screen "BWT Digital Inputs" 1280x800, template "Template"
   on GenerateScreen: "TitleUpdater"()
   TextField "Text field_37" at 16,52 size 263x26; Text 'BWT Control PLC (Rack 3)'
   TextField "Text field_38" at 16,122 size 55x22; Text 'I0.0'
   TextField "Text field_39" at 16,158 size 55x22; Text 'I0.1'
   TextField "Text field_40" at 16,194 size 55x22; Text 'I0.2'
   TextField "Text field_41" at 16,230 size 55x22; Text 'I0.3'
   TextField "Text field_42" at 16,265 size 55x22; Text 'I0.4'
   TextField "Text field_43" at 16,301 size 55x22; Text 'I0.5'
   TextField "Text field_44" at 16,337 size 55x22; Text 'I0.6'
   TextField "Text field_45" at 16,373 size 55x22; Text 'I0.7'
   Circle "Circle_33" at 76,122 size 20x20
      Appearance <- "10 DI_DATA_PS101"
   Circle "Circle_34" at 76,158 size 20x20
      Appearance <- "10 DI_DATA_E131_SHTDN"
   Circle "Circle_35" at 76,194 size 20x20
      Appearance <- "10 DI_DATA_R2_SPR_DI_0_2"
   Circle "Circle_36" at 76,230 size 20x20
      Appearance <- "10 DI_DATA_R2_SPR_DI_0_3"
   Circle "Circle_37" at 76,265 size 20x20
      Appearance <- "10 DI_DATA_X001_PWR_OK"
   Circle "Circle_38" at 76,301 size 20x20
      Appearance <- "10 DI_DATA_FD001_PWR_OK"
   Circle "Circle_39" at 76,337 size 20x20
      Appearance <- "10 DI_DATA_FD001_OK"
   Circle "Circle_40" at 76,373 size 20x20
      Appearance <- "103_Main_Burner_DB_DN_OK(1)"
   TextField "Text field_46" at 33,90 size 49x26; Text 'I0'
   TextField "Text field_47" at 16,441 size 55x22; Text 'I1.0'
   TextField "Text field_48" at 16,477 size 55x22; Text 'I1.1'
   TextField "Text field_49" at 16,513 size 55x22; Text 'I1.2'
   TextField "Text field_50" at 16,549 size 55x22; Text 'I1.3'
   TextField "Text field_51" at 16,584 size 55x22; Text 'I1.4'
   TextField "Text field_52" at 16,620 size 55x22; Text 'I1.5'
   TextField "Text field_53" at 16,656 size 55x22; Text 'I1.6'
   TextField "Text field_54" at 16,692 size 55x22; Text 'I1.7'
   Circle "Circle_41" at 76,441 size 20x20
      Appearance <- "10 DI_DATA_FS123"
   Circle "Circle_42" at 76,477 size 20x20
      Appearance <- "10 DI_DATA_FS115(1)"
   Circle "Circle_43" at 76,513 size 20x20
      Appearance <- "10 DI_DATA_FS320"
   Circle "Circle_44" at 76,549 size 20x20
      Appearance <- "10 DI_DATA_FS317"
   Circle "Circle_45" at 76,584 size 20x20
      Appearance <- "10 DI_DATA_P301_TRIPPED(1)"
   Circle "Circle_46" at 76,620 size 20x20
      Appearance <- "10 DI_DATA_P301_ENBLD"
   Circle "Circle_47" at 76,656 size 20x20
      Appearance <- "10 DI_DATA_R2_SPR_DI_1_6"
   Circle "Circle_48" at 76,692 size 20x20
      Appearance <- "10 DI_DATA_ESD_OK"
   TextField "Text field_55" at 33,409 size 49x26; Text 'I1'
   TextField "Text field_56" at 307,122 size 55x22; Text 'I2.0'
   TextField "Text field_57" at 307,158 size 55x22; Text 'I2.1'
   TextField "Text field_58" at 307,194 size 55x22; Text 'I2.2'
   TextField "Text field_59" at 307,230 size 55x22; Text 'I2.3'
   TextField "Text field_60" at 307,265 size 55x22; Text 'I2.4'
   TextField "Text field_61" at 307,301 size 55x22; Text 'I2.5'
   TextField "Text field_62" at 307,337 size 55x22; Text 'I2.6'
   TextField "Text field_63" at 307,373 size 55x22; Text 'I2.7'
   Circle "Circle_49" at 367,122 size 20x20
      Appearance <- "10 DI_DATA_E600_NOK"
   Circle "Circle_50" at 367,158 size 20x20
      Appearance <- "10 DI_DATA_E600_HIHI"
   Circle "Circle_51" at 367,194 size 20x20
      Appearance <- "10 DI_DATA_E600_LOLO"
   Circle "Circle_52" at 367,230 size 20x20
      Appearance <- "10 DI_DATA_E600_PWR_OK"
   Circle "Circle_53" at 367,265 size 20x20
      Appearance <- "10 DI_DATA_E700_PWR_OK"
   Circle "Circle_54" at 367,301 size 20x20
      Appearance <- "10 DI_DATA_E700_OPACITY"
   Circle "Circle_55" at 367,337 size 20x20
      Appearance <- "10 DI_DATA_TS403_FAULT(1)"
   Circle "Circle_56" at 367,373 size 20x20
      Appearance <- "10 DI_DATA_TS006"
   TextField "Text field_64" at 324,90 size 49x26; Text 'I2'
   TextField "Text field_65" at 305,441 size 46x22; Text 'I3.0'
   TextField "Text field_66" at 305,477 size 46x22; Text 'I3.1'
   TextField "Text field_67" at 305,513 size 46x22; Text 'I3.2'
   TextField "Text field_68" at 305,549 size 46x22; Text 'I3.3'
   TextField "Text field_69" at 305,584 size 46x22; Text 'I3.4'
   TextField "Text field_70" at 305,620 size 46x22; Text 'I3.5'
   TextField "Text field_71" at 305,656 size 46x22; Text 'I3.6'
   TextField "Text field_72" at 305,692 size 46x22; Text 'I3.7'
   Circle "Circle_57" at 365,441 size 20x20
      Appearance <- "10 DI_DATA_S2_8K1_OK"
   Circle "Circle_58" at 365,477 size 20x20
      Appearance <- "10 DI_DATA_E131_WRNG"
   Circle "Circle_59" at 365,513 size 20x20
      Appearance <- "10 DI_DATA_R2_SPR_DI_3_2"
   Circle "Circle_60" at 365,549 size 20x20
      Appearance <- "10 DI_DATA_E131_OK"
   Circle "Circle_61" at 365,584 size 20x20
      Appearance <- "10 DI_DATA_LS001"
   Circle "Circle_62" at 365,620 size 20x20
      Appearance <- "10 DI_DATA_P305_TRIPPED"
   Circle "Circle_63" at 365,656 size 20x20
      Appearance <- "10 DI_DATA_P305_ENBLD"
   Circle "Circle_64" at 365,692 size 20x20
      Appearance <- "10 DI_DATA_R2_SPR_DI_3_7"
   TextField "Text field_73" at 322,409 size 49x26; Text 'I3'
   Button "HmiScreenItemData_1" at 1,1 size 150x43; TextOn 'Back'; TextOff 'Commissioning'
      on Release: ActivateScreen("Commissioning Main Page", 0)
   TextField "Text field_107" at 105,111 size 243x23; Text 'CA Pressure Switch PS101'
   TextField "Text field_108" at 105,151 size 227x23; Text 'IA Comp Shutdown E131'
   TextField "Text field_109" at 104,191 size 112x23; Text 'Spare Input'
   TextField "Text field_110" at 104,225 size 112x23; Text 'Spare Input'
   TextField "Text field_111" at 104,257 size 258x23; Text 'Ignitor Power Healthy X001'
   TextField "Text field_112" at 104,292 size 181x42; Text 'FDU Power Healthy FD001'
   TextField "Text field_113" at 104,328 size 118x42; Text 'FDU Healthy FD001'
   TextField "Text field_114" at 104,365 size 215x42; Text 'Burner Flame Detected FD001'
   TextField "Text field_116" at 102,432 size 204x42; Text 'Pilot Ign. Air Flow Sw FS123'
   TextField "Text field_117" at 101,468 size 216x42; Text 'Main Atom Air Flow Sw FS115'
   TextField "Text field_118" at 101,504 size 182x42; Text 'Nozzle CW Flow Sw FS320'
   TextField "Text field_119" at 102,541 size 180x42; Text 'Jacket CW Flow Sw FS317'
   TextField "Text field_120" at 102,576 size 178x42; Text 'CSW Pump Tripped P301'
   TextField "Text field_121" at 105,611 size 180x42; Text 'CSW Pump Enabled P301'
   TextField "Text field_122" at 103,690 size 136x23; Text 'Ext. Shutdown'
   TextField "Text field_123" at 395,113 size 140x42; Text 'O2 System Fail E600'
   TextField "Text field_124" at 395,150 size 80x42; Text 'O2 Hi Hi E600'
   TextField "Text field_125" at 394,186 size 84x42; Text 'O2 Lo Lo E600'
   TextField "Text field_126" at 394,222 size 240x42; Text 'O2 System Power Healthy E600'
   TextField "Text field_127" at 394,256 size 257x42; Text 'Soot System Power Healthy E700'
   TextField "Text field_128" at 394,291 size 192x42; Text 'Soot System Opacity E700'
   TextField "Text field_129" at 394,328 size 199x42; Text 'IG Temp Hi Hi Switch TS403'
   TextField "Text field_130" at 395,366 size 225x42; Text 'IG Shell Temp Hi Switch TS006'
   TextField "Text field_131" at 394,437 size 181x23; Text 'IGG E-Stop Healthy'
   TextField "Text field_132" at 394,468 size 164x42; Text 'IA Comp Warning E131'
   TextField "Text field_133" at 393,509 size 112x23; Text 'Spare Input'
   TextField "Text field_134" at 393,611 size 248x42; Text 'Fresh Water Pump Tripped P305'
   TextField "Text field_135" at 393,648 size 250x42; Text 'Fresh Water Pump Enabled P305'
   TextField "Text field_136" at 394,688 size 112x23; Text 'Spare Input'
   TextField "Text field_137" at 395,540 size 159x42; Text 'IA Comp Healthy E131'
   TextField "Text field_138" at 394,576 size 222x42; Text 'Shell CW Level Hi Hi Sw LS001'
   TextField "Text field_115" at 105,654 size 112x23; Text 'Spare Input'
   AlarmView "Alarm view_1" at 0,777 size 1280x23
   TextField "Text field_1" at 23,309 size 1188x123; Text 'Re - Work Required Througout This page'
   Group "Group" at 455,41 size 373x50
   Button "HmiScreenItemData_8" at 469,45 size 355x40; TextOn 'Back'; TextOff 'Text'
   TextField "Screen title" at 455,41 size 373x50; Text 'Screen title'

screen "RIO 01 Digital Inputs" 1280x800, template "Template"
   on GenerateScreen: "TitleUpdater"()
   TextField "Text field_37" at 16,52 size 476x26; Text 'RIO #1 (Remote Inputs & Outputs Panel No. 1)'
   TextField "Text field_38" at 16,122 size 55x22; Text 'I0.0'
   TextField "Text field_39" at 16,157 size 55x22; Text 'I0.1'
   TextField "Text field_40" at 16,193 size 55x22; Text 'I0.2'
   TextField "Text field_41" at 16,229 size 55x22; Text 'I0.3'
   TextField "Text field_42" at 16,265 size 55x22; Text 'I0.4'
   TextField "Text field_43" at 16,301 size 55x22; Text 'I0.5'
   TextField "Text field_44" at 16,337 size 55x22; Text 'I0.6'
   TextField "Text field_45" at 16,373 size 55x22; Text 'I0.7'
   Circle "Circle_33" at 76,123 size 20x20
      Appearance <- "FPT GTT Isolation Valve Feedback - Opened"
   Circle "Circle_34" at 76,158 size 20x20
      Appearance <- "FPT GTT Isolation Valve Feedback - Closed"
   Circle "Circle_35" at 76,194 size 20x20
      Appearance <- "FPT Tank Vent Valve 1 Feedback - Opened"
   Circle "Circle_36" at 76,230 size 20x20
      Appearance <- "FPT Tank Vent Valve 1 Feedback - Closed"
   Circle "Circle_37" at 76,265 size 20x20
      Appearance <- "FPT Tank Vent Valve 2 Feedback - Opened"
   Circle "Circle_38" at 76,301 size 20x20
      Appearance <- "FPT Tank Vent Valve 2 Feedback - Closed"
   Circle "Circle_39" at 76,337 size 20x20
      Appearance <- "RIO1_SPR_DI_0_6"
   Circle "Circle_40" at 76,373 size 20x20
      Appearance <- "RIO1_SPR_DI_0_7"
   TextField "Text field_46" at 33,90 size 49x26; Text 'I0'
   TextField "Text field_47" at 16,441 size 55x22; Text 'I3.0'
   TextField "Text field_48" at 16,476 size 55x22; Text 'I3.1'
   TextField "Text field_49" at 16,512 size 55x22; Text 'I3.2'
   TextField "Text field_50" at 16,548 size 55x22; Text 'I3.3'
   TextField "Text field_51" at 16,584 size 55x22; Text 'I3.4'
   TextField "Text field_52" at 16,620 size 55x22; Text 'I3.5'
   TextField "Text field_53" at 16,656 size 55x22; Text 'I3.6'
   TextField "Text field_54" at 16,692 size 55x22; Text 'I3.7'
   Circle "Circle_41" at 76,442 size 20x20
      Appearance <- "Tank 1P GTT Isolation Valve Feedback - Opened"
   Circle "Circle_42" at 76,477 size 20x20
      Appearance <- "Tank 1P GTT Isolation Valve Feedback - Closed"
   Circle "Circle_43" at 76,513 size 20x20
      Appearance <- "Tank 1P Tank Vent Valve 1 Feedback - Opened"
   Circle "Circle_44" at 76,549 size 20x20
      Appearance <- "Tank 1P Tank Vent Valve 1 Feedback - Closed"
   Circle "Circle_45" at 76,585 size 20x20
      Appearance <- "Tank 1P Tank Vent Valve 2 Feedback - Opened"
   Circle "Circle_46" at 76,621 size 20x20
      Appearance <- "Tank 1P Tank Vent Valve 2 Feedback - Closed"
   Circle "Circle_47" at 76,657 size 20x20
      Appearance <- "RIO1_SPR_DI_3_6"
   Circle "Circle_48" at 76,693 size 20x20
      Appearance <- "RIO1_SPR_DI_3_7"
   TextField "Text field_55" at 33,409 size 49x26; Text 'I1'
   TextField "Text field_56" at 548,122 size 55x22; Text 'I6.0'
   TextField "Text field_57" at 548,157 size 55x22; Text 'I6.1'
   TextField "Text field_58" at 548,193 size 55x22; Text 'I6.2'
   TextField "Text field_59" at 548,229 size 55x22; Text 'I6.3'
   TextField "Text field_60" at 548,265 size 55x22; Text 'I6.4'
   TextField "Text field_61" at 548,301 size 55x22; Text 'I6.5'
   TextField "Text field_62" at 548,337 size 55x22; Text 'I6.6'
   TextField "Text field_63" at 548,373 size 55x22; Text 'I6.7'
   Circle "Circle_49" at 608,122 size 20x20
      Appearance <- "Tank 1S GTT Isolation Valve Feedback - Opened"
   Circle "Circle_50" at 608,157 size 20x20
      Appearance <- "Tank 1S GTT Isolation Valve Feedback - Closed"
   Circle "Circle_51" at 608,193 size 20x20
      Appearance <- "Tank 1S Tank Vent Valve 1 Feedback - Opened"
   Circle "Circle_52" at 608,229 size 20x20
      Appearance <- "Tank 1S Tank Vent Valve 1 Feedback - Closed"
   Circle "Circle_53" at 608,265 size 20x20
      Appearance <- "Tank 1S Tank Vent Valve 2 Feedback - Opened"
   Circle "Circle_54" at 608,301 size 20x20
      Appearance <- "Tank 1S Tank Vent Valve 2 Feedback - Closed"
   Circle "Circle_55" at 608,337 size 20x20
      Appearance <- "RIO1_SPR_DI_6_6"
   Circle "Circle_56" at 608,373 size 20x20
      Appearance <- "RIO1_SPR_DI_6_7"
   TextField "Text field_64" at 570,90 size 49x26; Text 'I2'
   TextField "Text field_65" at 546,441 size 46x22; Text 'I9.0'
   TextField "Text field_66" at 546,476 size 46x22; Text 'I9.1'
   TextField "Text field_67" at 546,512 size 46x22; Text 'I9.2'
   TextField "Text field_68" at 546,548 size 46x22; Text 'I9.3'
   TextField "Text field_69" at 546,584 size 46x22; Text 'I9.4'
   TextField "Text field_70" at 546,620 size 46x22; Text 'I9.5'
   TextField "Text field_71" at 546,656 size 46x22; Text 'I9.6'
   TextField "Text field_72" at 546,692 size 46x22; Text 'I9.7'
   Circle "Circle_57" at 606,441 size 20x20
      Appearance <- "FPT BWT Level High High Switch"
   Circle "Circle_58" at 606,476 size 20x20
      Appearance <- "RIO1 Tanks Pressure Switch Hi Hi"
   Circle "Circle_59" at 606,512 size 20x20
      Appearance <- "Tank 1P BWT Level High High Switch"
   Circle "Circle_60" at 606,548 size 20x20
      Appearance <- "Tank 1S BWT Level High High Switch"
   Circle "Circle_61" at 606,584 size 20x20
      Appearance <- "RIO1_SPR_DI_9_4"
   Circle "Circle_62" at 606,620 size 20x20
      Appearance <- "RIO1_SPR_DI_9_5"
   Circle "Circle_63" at 606,656 size 20x20
      Appearance <- "RIO1_SPR_DI_9_6"
   Circle "Circle_64" at 606,692 size 20x20
      Appearance <- "RIO1_SPR_DI_9_7"
   TextField "Text field_73" at 563,409 size 49x26; Text 'I3'
   Button "HmiScreenItemData_1" at 1,1 size 150x43; TextOn 'Back'; TextOff 'Commissioning'
      on Release: ActivateScreen("Commissioning Main Page", 0)
   TextField "Text field_107" at 105,114 size 348x38; Text 'FPT GTT Isolation Valve Feedback - Opened CV422'
   TextField "Text field_108" at 105,149 size 340x38; Text 'FPT GTT Isolation Valve Feedback - Closed CV422'
   TextField "Text field_109" at 105,184 size 337x38; Text 'FPT Tank Vent Valve 1 Feedback - Opened CV441-FPTA'
   TextField "Text field_110" at 105,220 size 329x38; Text 'FPT Tank Vent Valve 1 Feedback - Closed CV441-FPTA'
   TextField "Text field_111" at 105,255 size 337x38; Text 'FPT Tank Vent Valve 2 Feedback - Opened CV441-FPTB'
   TextField "Text field_112" at 105,291 size 329x38; Text 'FPT Tank Vent Valve 2 Feedback - Closed CV441-FPTB'
   TextField "Text field_113" at 104,328 size 100x21; Text 'Spare Input'
   TextField "Text field_114" at 104,365 size 100x21; Text 'Spare Input'
   TextField "Text field_116" at 102,429 size 382x38; Text 'Tank 1P GTT Isolation Valve Feedback - Opened CV422'
   TextField "Text field_117" at 102,465 size 374x38; Text 'Tank 1P GTT Isolation Valve Feedback - Closed CV422'
   TextField "Text field_118" at 102,501 size 371x38; Text 'Tank 1P Tank Vent Valve 1 Feedback - Opened CV441-1PA'
   TextField "Text field_119" at 102,537 size 363x38; Text 'Tank 1P Tank Vent Valve 1 Feedback - Closed CV441-1PA'
   TextField "Text field_120" at 102,573 size 371x38; Text 'Tank 1P Tank Vent Valve 2 Feedback - Opened CV441-1PB'
   TextField "Text field_121" at 102,609 size 363x38; Text 'Tank 1P Tank Vent Valve 2 Feedback - Closed CV441-1PB'
   TextField "Text field_122" at 102,690 size 100x21; Text 'Spare Input'
   TextField "Text field_123" at 636,113 size 382x38; Text 'Tank 1S GTT Isolation Valve Feedback - Opened CV421'
   TextField "Text field_124" at 636,148 size 374x38; Text 'Tank 1S GTT Isolation Valve Feedback - Closed CV421'
   TextField "Text field_125" at 636,184 size 371x38; Text 'Tank 1S Tank Vent Valve 1 Feedback - Opened CV440-1SA'
   TextField "Text field_126" at 636,219 size 363x38; Text 'Tank 1S Tank Vent Valve 1 Feedback - Closed CV440-1SA'
   TextField "Text field_127" at 636,255 size 371x38; Text 'Tank 1S Tank Vent Valve 2 Feedback - Opened CV440-1SB'
   TextField "Text field_128" at 636,291 size 363x38; Text 'Tank 1S Tank Vent Valve 2 Feedback - Closed CV440-1SB'
   TextField "Text field_129" at 636,328 size 100x21; Text 'Spare Input'
   TextField "Text field_130" at 636,366 size 100x21; Text 'Spare Input'
   TextField "Text field_131" at 635,431 size 260x38; Text 'FPT BWT Level High High Switch LS425-FPT'
   TextField "Text field_132" at 635,467 size 270x38; Text 'RIO1 Tanks Pressure Switch Hi Hi PS436-FPT/1P/1S'
   TextField "Text field_133" at 635,503 size 294x38; Text 'Tank 1P BWT Level High High Switch LS425-1P'
   TextField "Text field_134" at 635,611 size 100x21; Text 'Spare Input'
   TextField "Text field_135" at 635,648 size 100x21; Text 'Spare Input'
   TextField "Text field_136" at 635,688 size 100x21; Text 'Spare Input'
   TextField "Text field_137" at 635,539 size 294x38; Text 'Tank 1S BWT Level High High Switch LS425-1S'
   TextField "Text field_138" at 635,576 size 100x21; Text 'Spare Input'
   TextField "Text field_115" at 102,654 size 100x21; Text 'Spare Input'
   AlarmView "Alarm view_1" at 0,777 size 1280x23
   Group "Group" at 455,41 size 373x50
   Button "HmiScreenItemData_8" at 469,45 size 355x40; TextOn 'Back'; TextOff 'Text'
      on Click: "TitleUpdater"()
   TextField "Screen title" at 455,41 size 373x50; Text 'Screen title'

screen "IGG Digital Outputs" 1280x800, template "Template"
   on GenerateScreen: "TitleUpdater"()
   Button "HmiScreenItemData_1" at 1,1 size 150x43; TextOn 'Back'; TextOff 'Commissioning'
      on Release: ActivateScreen("Commissioning Main Page", 0)
   AlarmView "Alarm view_1" at 0,777 size 1280x23
   TextField "Text field_1" at 395,239 size 55x22; Text 'Q0.0'
   TextField "Text field_2" at 395,290 size 55x22; Text 'Q0.1'
   TextField "Text field_3" at 395,342 size 55x22; Text 'Q0.2'
   TextField "Text field_4" at 395,394 size 55x22; Text 'Q0.3'
   TextField "Text field_5" at 395,446 size 55x22; Text 'Q0.4'
   TextField "Text field_6" at 395,498 size 55x22; Text 'Q0.5'
   TextField "Text field_7" at 395,550 size 55x22; Text 'Q0.6'
   TextField "Text field_8" at 395,602 size 55x22; Text 'Q0.7'
   Circle "Circle_1" at 455,239 size 20x20
      Appearance <- "14_DQ_Data_E500A_CNTRL"
   Circle "Circle_2" at 455,290 size 20x20
      Appearance <- "14_DQ_Data_E500B_CNTRL"
   Circle "Circle_3" at 455,342 size 20x20
      Appearance <- "14_DQ_Data_E139_CNTRL"
   Circle "Circle_4" at 455,394 size 20x20
      Appearance <- "14_DQ_Data_CV311_312_CNTRL"
   Circle "Circle_5" at 455,446 size 20x20
      Appearance <- "14_DQ_Data_CV321_322_CNTRL"
   Circle "Circle_6" at 455,498 size 20x20
      Appearance <- "14_DQ_Data_CV401_CNTRL"
   Circle "Circle_7" at 455,550 size 20x20
      Appearance <- "14_DQ_Data_CV431_432_CNTRL"
   Circle "Circle_8" at 455,602 size 20x20
      Appearance <- "14_DQ_Data_R2_SPR_DQ_0_7"
   TextField "Text field_9" at 412,206 size 49x26; Text 'Q0'
   TextField "Text field_10" at 698,239 size 55x22; Text 'Q1.0'
   TextField "Text field_11" at 698,290 size 55x22; Text 'Q1.1'
   TextField "Text field_12" at 698,342 size 55x22; Text 'Q1.2'
   TextField "Text field_13" at 698,394 size 55x22; Text 'Q1.3'
   TextField "Text field_14" at 698,446 size 55x22; Text 'Q1.4'
   TextField "Text field_15" at 698,498 size 55x22; Text 'Q1.5'
   TextField "Text field_16" at 698,550 size 55x22; Text 'Q1.6'
   TextField "Text field_17" at 698,602 size 55x22; Text 'Q1.7'
   Circle "Circle_9" at 758,239 size 20x20
      Appearance <- "14_DQ_Data_R2_SPR_DQ_1_0"
   Circle "Circle_10" at 758,290 size 20x20
      Appearance <- "14_DQ_Data_24K2"
   Circle "Circle_11" at 758,342 size 20x20
      Appearance <- "14_DQ_Data_24K3"
   Circle "Circle_12" at 758,394 size 20x20
      Appearance <- "14_DQ_Data_24K4"
   Circle "Circle_13" at 758,446 size 20x20
      Appearance <- "14_DQ_Data_24PF1"
   Circle "Circle_14" at 758,498 size 20x20
      Appearance <- "14_DQ_Data_24PF2"
   Circle "Circle_15" at 758,550 size 20x20
      Appearance <- "14_DQ_Data_24PF3"
   Circle "Circle_16" at 758,602 size 20x20
      Appearance <- "14_DQ_Data_24PF4"
   TextField "Text field_18" at 715,206 size 49x26; Text 'Q1'
   TextField "Text field_37" at 328,167 size 254x26; Text 'IGG System PLC (Rack 1)'
   Button "Button_9" at 330,493 size 60x35; TextOff 'Override'
      on Press: InvertBit("80_From_HMI_MAN_DQ_0_5")
      Visibility <- "82_To_HMI_CRNT_MODE_IGG"
   Button "Button_10" at 330,441 size 60x35; TextOff 'Override'
      on Press: InvertBit("80_From_HMI_MAN_DQ_0_4")
      Visibility <- "82_To_HMI_CRNT_MODE_IGG"
   Button "Button_11" at 330,388 size 60x35; TextOff 'Override'
      on Press: InvertBit("80_From_HMI_MAN_DQ_0_3")
      Visibility <- "82_To_HMI_CRNT_MODE_IGG"
   Button "Button_12" at 631,596 size 60x35; TextOff 'Override'
      on Press: InvertBit("80_From_HMI_MAN_DQ_1_7")
      Visibility <- "82_To_HMI_CRNT_MODE_IGG"
   Button "Button_14" at 631,283 size 60x35; TextOff 'Override'
      on Press: InvertBit("80_From_HMI_MAN_DQ_1_1")
      Visibility <- "82_To_HMI_CRNT_MODE_IGG"
   TextField "Text field_56" at 481,239 size 140x22; Text 'Fuel Pump 1 E500A'
   TextField "Text field_57" at 481,290 size 140x22; Text 'Fuel Pump 2 E500B'
   TextField "Text field_58" at 481,342 size 140x22; Text 'CA Blower E139'
   TextField "Text field_59" at 481,394 size 140x22; Text 'CSW Inlet Valves CV311'
   TextField "Text field_60" at 481,446 size 140x22; Text 'CSW Drain Valves CV322'
   TextField "Text field_61" at 481,498 size 140x22; Text 'IG Supply Valve CV401'
   TextField "Text field_62" at 481,549 size 140x22; Text 'CB/BWTS Valve CV432'
   TextField "Text field_63" at 481,602 size 140x22; Text 'Spare Output'
   TextField "Text field_64" at 786,242 size 140x22; Text 'Spare Output'
   TextField "Text field_65" at 786,290 size 140x22; Text 'Atmospheric Alarm'
   TextField "Text field_66" at 786,342 size 140x22; Text 'IGG Shutdown Alarm'
   TextField "Text field_67" at 786,394 size 140x22; Text 'IGG Warning Alarm'
   TextField "Text field_68" at 786,446 size 140x22; Text 'IGG Running'
   TextField "Text field_69" at 786,497 size 140x22; Text 'Shutdown Alarm'
   TextField "Text field_70" at 786,550 size 140x22; Text 'Warning Alarm'
   TextField "Text field_71" at 786,602 size 140x22; Text 'Buzzer'
   Button "Button_15" at 330,336 size 60x35; TextOff 'Override'
      on Press: InvertBit("80_From_HMI_MAN_DQ_0_2")
      Visibility <- "82_To_HMI_CRNT_MODE_IGG"
   Button "Button_16" at 330,283 size 60x35; TextOff 'Override'
      on Press: InvertBit("80_From_HMI_MAN_DQ_0_1")
      Visibility <- "82_To_HMI_CRNT_MODE_IGG"
   Button "Button_17" at 330,546 size 60x35; TextOff 'Override'
      on Press: InvertBit("80_From_HMI_MAN_DQ_0_6")
      Visibility <- "82_To_HMI_CRNT_MODE_IGG"
   Button "Button_18" at 330,599 size 60x35; TextOff 'Override'
      on Press: InvertBit("80_From_HMI_MAN_DQ_0_7(1)")
      Visibility <- "82_To_HMI_CRNT_MODE_IGG"
   Button "Button_19" at 330,231 size 60x35; TextOff 'Override'
      on Press: InvertBit("80_From_HMI_MAN_DQ_0_0")
      Visibility <- "82_To_HMI_CRNT_MODE_IGG"
   Button "Button_20" at 631,231 size 60x35; TextOff 'Override'
      on Press: InvertBit("80_From_HMI_MAN_DQ_1_0(1)")
      Visibility <- "82_To_HMI_CRNT_MODE_IGG"
   Button "Button_21" at 631,335 size 60x35; TextOff 'Override'
      on Press: InvertBit("80_From_HMI_MAN_DQ_1_2")
      Visibility <- "82_To_HMI_CRNT_MODE_IGG"
   Button "Button_22" at 631,387 size 60x35; TextOff 'Override'
      on Press: InvertBit("80_From_HMI_MAN_DQ_1_3")
      Visibility <- "82_To_HMI_CRNT_MODE_IGG"
   Button "Button_23" at 631,439 size 60x35; TextOff 'Override'
      on Press: InvertBit("80_From_HMI_MAN_DQ_1_4")
      Visibility <- "82_To_HMI_CRNT_MODE_IGG"
   Button "Button_24" at 631,491 size 60x35; TextOff 'Override'
      on Press: InvertBit("80_From_HMI_MAN_DQ_1_5")
      Visibility <- "82_To_HMI_CRNT_MODE_IGG"
   Button "Button_25" at 631,543 size 60x35; TextOff 'Override'
      on Press: InvertBit("80_From_HMI_MAN_DQ_1_6(1)")
      Visibility <- "82_To_HMI_CRNT_MODE_IGG"
   Group "Group" at 455,41 size 373x50
   Button "HmiScreenItemData_8" at 469,45 size 355x40; TextOn 'Back'; TextOff 'Text'
   TextField "Screen title" at 455,41 size 373x50; Text 'Screen title'

screen "BWT Digital Outputs" 1280x800, template "Template"
   on GenerateScreen: "TitleUpdater"()
   TextField "Text field_1" at 79,178 size 55x22; Text 'Q0.0'
   TextField "Text field_2" at 79,229 size 55x22; Text 'Q0.1'
   TextField "Text field_3" at 79,281 size 55x22; Text 'Q0.2'
   TextField "Text field_4" at 79,333 size 55x22; Text 'Q0.3'
   TextField "Text field_5" at 79,385 size 55x22; Text 'Q0.4'
   TextField "Text field_6" at 79,437 size 55x22; Text 'Q0.5'
   TextField "Text field_7" at 79,489 size 55x22; Text 'Q0.6'
   TextField "Text field_8" at 79,541 size 55x22; Text 'Q0.7'
   Circle "Circle_1" at 139,178 size 20x20
      Appearance <- "14_DQ_Data_E500A_CNTRL"
   Circle "Circle_2" at 139,229 size 20x20
      Appearance <- "14_DQ_Data_E500B_CNTRL"
   Circle "Circle_3" at 139,281 size 20x20
      Appearance <- "14_DQ_Data_E139_CNTRL"
   Circle "Circle_4" at 139,333 size 20x20
      Appearance <- "14_DQ_Data_CV311_312_CNTRL"
   Circle "Circle_5" at 139,385 size 20x20
      Appearance <- "14_DQ_Data_CV321_322_CNTRL"
   Circle "Circle_6" at 139,437 size 20x20
      Appearance <- "14_DQ_Data_CV401_CNTRL"
   Circle "Circle_7" at 139,489 size 20x20
      Appearance <- "14_DQ_Data_CV431_432_CNTRL"
   Circle "Circle_8" at 139,541 size 20x20
      Appearance <- "14_DQ_Data_R2_SPR_DQ_0_7"
   TextField "Text field_9" at 96,145 size 49x26; Text 'Q0'
   TextField "Text field_10" at 382,178 size 55x22; Text 'Q1.0'
   TextField "Text field_11" at 382,229 size 55x22; Text 'Q1.1'
   TextField "Text field_12" at 382,281 size 55x22; Text 'Q1.2'
   TextField "Text field_13" at 382,333 size 55x22; Text 'Q1.3'
   TextField "Text field_14" at 382,385 size 55x22; Text 'Q1.4'
   TextField "Text field_15" at 382,437 size 55x22; Text 'Q1.5'
   TextField "Text field_16" at 382,489 size 55x22; Text 'Q1.6'
   TextField "Text field_17" at 382,541 size 55x22; Text 'Q1.7'
   Circle "Circle_9" at 442,178 size 20x20
      Appearance <- "14_DQ_Data_R2_SPR_DQ_1_0"
   Circle "Circle_10" at 442,229 size 20x20
      Appearance <- "14_DQ_Data_24K2"
   Circle "Circle_11" at 442,281 size 20x20
      Appearance <- "14_DQ_Data_24K3"
   Circle "Circle_12" at 442,333 size 20x20
      Appearance <- "14_DQ_Data_24K4"
   Circle "Circle_13" at 442,385 size 20x20
      Appearance <- "14_DQ_Data_24PF1"
   Circle "Circle_14" at 442,437 size 20x20
      Appearance <- "14_DQ_Data_24PF2"
   Circle "Circle_15" at 442,489 size 20x20
      Appearance <- "14_DQ_Data_24PF3"
   Circle "Circle_16" at 442,541 size 20x20
      Appearance <- "14_DQ_Data_24PF4"
   TextField "Text field_18" at 399,145 size 49x26; Text 'Q1'
   TextField "Text field_37" at 12,106 size 263x26; Text 'BWT Control PLC (Rack 3)'
   Button "HmiScreenItemData_1" at 1,1 size 150x43; TextOn 'Back'; TextOff 'Commissioning'
      on Release: ActivateScreen("Commissioning Main Page", 0)
   Button "Button_9" at 14,432 size 60x35; TextOff 'Override'
      on Press: InvertBit("80_From_HMI_MAN_DQ_0_5")
      Visibility <- "82_To_HMI_CRNT_MODE_IGG"
   Button "Button_10" at 14,380 size 60x35; TextOff 'Override'
      on Press: InvertBit("80_From_HMI_MAN_DQ_0_4")
      Visibility <- "82_To_HMI_CRNT_MODE_IGG"
   Button "Button_11" at 14,327 size 60x35; TextOff 'Override'
      on Press: InvertBit("80_From_HMI_MAN_DQ_0_3")
      Visibility <- "82_To_HMI_CRNT_MODE_IGG"
   Button "Button_12" at 315,535 size 60x35; TextOff 'Override'
      on Press: InvertBit("80_From_HMI_MAN_DQ_1_7")
      Visibility <- "82_To_HMI_CRNT_MODE_IGG"
   Button "Button_14" at 315,222 size 60x35; TextOff 'Override'
      on Press: InvertBit("80_From_HMI_MAN_DQ_1_1")
      Visibility <- "82_To_HMI_CRNT_MODE_IGG"
   TextField "Text field_56" at 165,174 size 117x42; Text 'Fuel Pump 1 E500A'
   TextField "Text field_57" at 165,223 size 117x42; Text 'Fuel Pump 2 E500B'
   TextField "Text field_58" at 165,277 size 100x42; Text 'CA Blower E139'
   TextField "Text field_59" at 165,327 size 161x42; Text 'CSW Inlet Valves CV311'
   TextField "Text field_60" at 165,378 size 166x42; Text 'CSW Drain Valves CV322'
   TextField "Text field_61" at 165,434 size 149x42; Text 'IG Supply Valve CV401'
   TextField "Text field_62" at 165,489 size 154x42; Text 'CB/BWTS Valve CV432'
   TextField "Text field_63" at 165,538 size 125x23; Text 'Spare Output'
   TextField "Text field_64" at 470,175 size 125x23; Text 'Spare Output'
   TextField "Text field_65" at 470,224 size 178x23; Text 'Atmospheric Alarm'
   TextField "Text field_66" at 470,278 size 194x23; Text 'IGG Shutdown Alarm'
   TextField "Text field_67" at 470,328 size 180x23; Text 'IGG Warning Alarm'
   TextField "Text field_68" at 470,379 size 119x23; Text 'IGG Running'
   TextField "Text field_69" at 470,431 size 154x23; Text 'Shutdown Alarm'
   TextField "Text field_70" at 470,490 size 140x23; Text 'Warning Alarm'
   TextField "Text field_71" at 470,539 size 67x23; Text 'Buzzer'
   Button "Button_15" at 14,275 size 60x35; TextOff 'Override'
      on Press: InvertBit("80_From_HMI_MAN_DQ_0_2")
      Visibility <- "82_To_HMI_CRNT_MODE_IGG"
   Button "Button_16" at 14,222 size 60x35; TextOff 'Override'
      on Press: InvertBit("80_From_HMI_MAN_DQ_0_1")
      Visibility <- "82_To_HMI_CRNT_MODE_IGG"
   Button "Button_17" at 14,485 size 60x35; TextOff 'Override'
      on Press: InvertBit("80_From_HMI_MAN_DQ_0_6")
      Visibility <- "82_To_HMI_CRNT_MODE_IGG"
   Button "Button_18" at 14,538 size 60x35; TextOff 'Override'
      on Press: InvertBit("80_From_HMI_MAN_DQ_0_7(1)")
      Visibility <- "82_To_HMI_CRNT_MODE_IGG"
   Button "Button_19" at 14,170 size 60x35; TextOff 'Override'
      on Press: InvertBit("80_From_HMI_MAN_DQ_0_0")
      Visibility <- "82_To_HMI_CRNT_MODE_IGG"
   Button "Button_20" at 315,170 size 60x35; TextOff 'Override'
      on Press: InvertBit("80_From_HMI_MAN_DQ_1_0(1)")
      Visibility <- "82_To_HMI_CRNT_MODE_IGG"
   Button "Button_21" at 315,274 size 60x35; TextOff 'Override'
      on Press: InvertBit("80_From_HMI_MAN_DQ_1_2")
      Visibility <- "82_To_HMI_CRNT_MODE_IGG"
   Button "Button_22" at 315,326 size 60x35; TextOff 'Override'
      on Press: InvertBit("80_From_HMI_MAN_DQ_1_3")
      Visibility <- "82_To_HMI_CRNT_MODE_IGG"
   Button "Button_23" at 315,378 size 60x35; TextOff 'Override'
      on Press: InvertBit("80_From_HMI_MAN_DQ_1_4")
      Visibility <- "82_To_HMI_CRNT_MODE_IGG"
   Button "Button_24" at 315,430 size 60x35; TextOff 'Override'
      on Press: InvertBit("80_From_HMI_MAN_DQ_1_5")
      Visibility <- "82_To_HMI_CRNT_MODE_IGG"
   Button "Button_25" at 315,482 size 60x35; TextOff 'Override'
      on Press: InvertBit("80_From_HMI_MAN_DQ_1_6(1)")
      Visibility <- "82_To_HMI_CRNT_MODE_IGG"
   AlarmView "Alarm view_1" at 0,777 size 1280x23
   TextField "Text field_19" at 23,309 size 1188x123; Text 'Re - Work Required Througout This page'
   Group "Group" at 455,41 size 373x50
   Button "HmiScreenItemData_8" at 469,45 size 355x40; TextOn 'Back'; TextOff 'Text'
   TextField "Screen title" at 455,41 size 373x50; Text 'Screen title'

screen "BWT Analogue Inputs" 1280x800, template "Template"
   on GenerateScreen: "TitleUpdater"()
   IOField "I/O field_62" at 1208,191 size 60x22; FormatPattern 99.9
   IOField "I/O field_61" at 1140,191 size 60x22; FormatPattern 99.9
   Button "HmiScreenItemData_1" at 1,1 size 150x43; TextOn 'Back'; TextOff 'Commissioning'
      on Release: ActivateScreen("Commissioning Main Page", 0)
   TextField "Text field_82" at 60,150 size 220x22; Text 'PIT-102 - CA Pressure (Pre-Ignition)'
   TextField "Text field_90" at 286,124 size 64x20; Text 'Reading'
   IOField "I/O field_2" at 287,150 size 70x22; FormatPattern 9999; Unit  mBar
      ProcessValue <- "12_AI_Data_PIT102_SCALED(1)"
   TextField "Text field_1" at 359,124 size 68x20; Text 'Low Low'
   IOField "I/O field_1" at 361,150 size 60x22; Authorization "Parameter Change"; FormatPattern 9999
      ProcessValue <- "84_Setpoints_PIT102_Pilot_LowLow"
   TextField "Text field_2" at 442,124 size 37x20; Text 'Low'
   IOField "I/O field_3" at 429,150 size 60x22; Authorization "Parameter Change"; FormatPattern 9999
      ProcessValue <- "84_Setpoints_PIT102_Pilot_Low"
   TextField "Text field_3" at 509,124 size 37x20; Text 'High'
   IOField "I/O field_4" at 497,150 size 60x22; Authorization "Parameter Change"; FormatPattern 9999
      ProcessValue <- "84_Setpoints_PIT102_Pilot_High"
   TextField "Text field_4" at 561,124 size 74x20; Text 'High High'
   IOField "I/O field_5" at 565,150 size 60x22; Authorization "Parameter Change"; FormatPattern 9999
      ProcessValue <- "84_Setpoints_PIT102_Pilot_HighHigh"
   TextField "Text field_5" at 434,100 size 76x20; Text 'Setpoints'
   TextField "Text field_6" at 7,150 size 53x22; Text 'IW112'
   TextField "Text field_7" at 60,270 size 220x22; Text 'TIT-401 - IG Temperature'
   IOField "I/O field_6" at 287,270 size 70x22; FormatPattern s999.9; Unit  °C
      ProcessValue <- "12_AI_Data_TIT401_SCALED"
   IOField "I/O field_7" at 361,270 size 60x22; FormatPattern s999.9
   IOField "I/O field_8" at 429,270 size 60x22; FormatPattern s999.9
   IOField "I/O field_9" at 497,270 size 60x22; Authorization "Parameter Change"; FormatPattern s999.9
      ProcessValue <- "84_Setpoints_TIT401_High"
   IOField "I/O field_10" at 565,270 size 60x22; Authorization "Parameter Change"; FormatPattern s999.9
      ProcessValue <- "84_Setpoints_TIT401_HighHigh"
   TextField "Text field_8" at 7,270 size 53x22; Text 'IW114'
   TextField "Text field_9" at 60,310 size 220x22; Text 'PIT-402 - IG Outlet Pres. (Pre-Ignitn.)'
   IOField "I/O field_11" at 287,310 size 70x22; FormatPattern 9999; Unit  mBar
      ProcessValue <- "12_AI_Data_PIT402_SCALED"
   IOField "I/O field_12" at 361,310 size 60x22; Authorization "Parameter Change"; FormatPattern 9999
      ProcessValue <- "84_Setpoints_PIT402_Pilot_LowLow"
   IOField "I/O field_13" at 429,310 size 60x22; Authorization "Parameter Change"; FormatPattern 9999
      ProcessValue <- "84_Setpoints_PIT402_Pilot_Low"
   IOField "I/O field_14" at 497,310 size 60x22; Authorization "Parameter Change"; FormatPattern 9999
      ProcessValue <- "84_Setpoints_PIT402_Pilot_High"
   IOField "I/O field_15" at 565,310 size 60x22; Authorization "Parameter Change"; FormatPattern 9999
      ProcessValue <- "84_Setpoints_PIT402_Pilot_HighHigh"
   TextField "Text field_10" at 7,310 size 53x22; Text 'IW116'
   TextField "Text field_11" at 60,430 size 220x22; Text 'CV-403 - IG Vent Valve Position Fbk'
   IOField "I/O field_16" at 287,430 size 70x22; FormatPattern 999; Unit  %
      ProcessValue <- "12_AI_Data_CV403_SCALED"
   IOField "I/O field_17" at 361,430 size 60x22; FormatPattern 999
   IOField "I/O field_18" at 429,430 size 60x22; FormatPattern 999
   IOField "I/O field_19" at 497,430 size 60x22; FormatPattern 999
   IOField "I/O field_20" at 565,430 size 60x22; FormatPattern 999
   TextField "Text field_12" at 7,430 size 53x22; Text 'IW118'
   TextField "Text field_13" at 60,470 size 220x22; Text 'CA Blower RPM'
   IOField "I/O field_21" at 287,470 size 70x22; FormatPattern 9999; Unit  RPM
      ProcessValue <- "12_AI_Data_E139_RPM_SCALED"
   IOField "I/O field_22" at 361,470 size 60x22; FormatPattern 9999
   IOField "I/O field_23" at 429,470 size 60x22; FormatPattern 9999
   IOField "I/O field_24" at 497,470 size 60x22; FormatPattern 9999
   IOField "I/O field_25" at 565,470 size 60x22; FormatPattern 9999
   TextField "Text field_14" at 7,470 size 54x22; Text 'IW120'
   TextField "Text field_15" at 61,511 size 220x22; Text 'CA Blower Current'
   IOField "I/O field_26" at 288,511 size 70x22; FormatPattern 999.9; Unit  A
      ProcessValue <- "12_AI_Data_E139_AMPS_SCALED"
   IOField "I/O field_27" at 362,511 size 60x22; FormatPattern 9999
   IOField "I/O field_28" at 430,511 size 60x22; FormatPattern 9999
   TextField "Text field_16" at 8,511 size 54x22; Text 'IW122'
   TextField "Text field_17" at 61,552 size 220x22; Text 'LIT-305 - FW Bulk Tank Level'
   IOField "I/O field_31" at 288,552 size 70x22; FormatPattern 99.9; Unit  %
      ProcessValue <- "12_AI_Data_LIT305_SCALED"
   TextField "Text field_18" at 8,552 size 53x22; Text 'IW124'
   TextField "Text field_19" at 61,592 size 220x22; Text 'Spare'
   IOField "I/O field_36" at 288,592 size 70x22; FormatPattern 9.9; Unit  
      ProcessValue <- "12_AI_Data_R1_SPR_AI_126_SCALED"
   IOField "I/O field_37" at 362,592 size 60x22; FormatPattern 9.9
   IOField "I/O field_38" at 430,592 size 60x22; FormatPattern 9.9
   IOField "I/O field_39" at 498,592 size 60x22; FormatPattern 9.9
   IOField "I/O field_40" at 566,592 size 60x22; FormatPattern 9.9
   TextField "Text field_20" at 8,592 size 53x22; Text 'IW126'
   TextField "Text field_21" at 703,151 size 220x22; Text 'Atmospheric Oxygen 1'
   IOField "I/O field_41" at 930,151 size 70x22; FormatPattern 99.99; Unit %
      ProcessValue <- "12_AI_Data_AT_O2_01_SCALED"
   IOField "I/O field_42" at 1004,151 size 60x22; Authorization "Commissioning"; FormatPattern 99.9
      ProcessValue <- "84_Setpoints_AT_O2_1_LowLow"
   IOField "I/O field_43" at 1072,151 size 60x22; Authorization "Commissioning"; FormatPattern 99.9
      ProcessValue <- "84_Setpoints_AT_O2_1_Low"
   IOField "I/O field_44" at 1140,151 size 60x22; FormatPattern 99.9
   IOField "I/O field_45" at 1208,151 size 60x22; FormatPattern 99.9
   TextField "Text field_22" at 650,151 size 53x22; Text 'IW128'
   TextField "Text field_23" at 703,191 size 220x22; Text 'Atmospheric Oxygen 2'
   IOField "I/O field_46" at 930,191 size 70x22; FormatPattern 99.99; Unit %
      ProcessValue <- "12_AI_Data_AT_O2_02_SCALED"
   TextField "Text field_24" at 650,191 size 53x22; Text 'IW130'
   TextField "Text field_26" at 928,124 size 64x20; Text 'Reading'
   TextField "Text field_27" at 1001,124 size 68x20; Text 'Low Low'
   TextField "Text field_28" at 1082,124 size 37x20; Text 'Low'
   TextField "Text field_29" at 1150,124 size 37x20; Text 'High'
   TextField "Text field_30" at 1203,124 size 74x20; Text 'High High'
   TextField "Text field_31" at 1076,100 size 76x20; Text 'Setpoints'
   TextField "Text field_51" at 703,231 size 220x22; Text 'Spare'
   IOField "I/O field_101" at 930,231 size 70x22; FormatPattern 99.9
      ProcessValue <- "12_AI_Data_R1_SPR_AI_132_SCALED"
   TextField "Text field_56" at 650,231 size 53x22; Text 'IW132'
   TextField "Text field_57" at 703,271 size 220x22; Text 'TIT-315 - Shell CSW Temperature'
   IOField "I/O field_106" at 930,271 size 70x22; FormatPattern s999.9; Unit  °C
      ProcessValue <- "12_AI_Data_TIT315_SCALED"
   IOField "I/O field_107" at 1004,271 size 60x22; FormatPattern s999.9
   IOField "I/O field_108" at 1072,271 size 60x22; FormatPattern s999.9
   TextField "Text field_58" at 650,271 size 54x22; Text 'IW134'
   TextField "Text field_59" at 703,311 size 220x22; Text 'TIT-319 - Inlet CSW Temperature'
   IOField "I/O field_111" at 930,311 size 70x22; FormatPattern s999.9; Unit  °C
      ProcessValue <- "12_AI_Data_TIT319_SCALED"
   IOField "I/O field_112" at 1004,311 size 60x22; FormatPattern s999.9
   IOField "I/O field_113" at 1072,311 size 60x22; FormatPattern s999.9
   TextField "Text field_60" at 650,311 size 53x22; Text 'IW136'
   TextField "Text field_61" at 703,351 size 220x22; Text 'TIT-360 - Outlet CSW Temperature'
   IOField "I/O field_116" at 930,351 size 70x22; FormatPattern s999.9; Unit  °C
      ProcessValue <- "12_AI_Data_TIT360_SCALED"
   IOField "I/O field_117" at 1004,351 size 60x22; FormatPattern s999.9
   IOField "I/O field_118" at 1072,351 size 60x22; FormatPattern s999.9
   TextField "Text field_62" at 650,351 size 53x22; Text 'IW138'
   TextField "Text field_63" at 703,391 size 220x22; Text 'PIT-359 - Inlet CSW Pressure'
   IOField "I/O field_121" at 930,391 size 70x22; FormatPattern 99.9; Unit  Bar
      ProcessValue <- "12_AI_Data_PIT359_SCALED"
   TextField "Text field_64" at 650,391 size 53x22; Text 'IW140'
   TextField "Text field_41" at 133,124 size 89x20; Text 'Description'
   TextField "Text field_42" at 771,124 size 89x20; Text 'Description'
   TextField "Text field_43" at 17,124 size 37x20; Text 'AI'
   TextField "Text field_44" at 661,124 size 37x20; Text 'AI'
   TextField "Text field_47" at 702,431 size 220x22; Text 'PIT-316 - Outlet CSW Pressure'
   IOField "I/O field_81" at 929,431 size 70x22; FormatPattern 99.9; Unit  Bar
      ProcessValue <- "12_AI_Data_PIT316_SCALED"
   TextField "Text field_48" at 649,431 size 53x22; Text 'IW142'
   IOField "I/O field_109" at 1140,271 size 60x22; Authorization "Parameter Change"; FormatPattern s999.9
      ProcessValue <- "84_Setpoints_TIT315_High"
   IOField "I/O field_110" at 1208,271 size 60x22; Authorization "Parameter Change"; FormatPattern s999.9
      ProcessValue <- "84_Setpoints_TIT315_HighHigh"
   IOField "I/O field_114" at 1140,311 size 60x22; Authorization "Parameter Change"; FormatPattern s999.9
      ProcessValue <- "84_Setpoints_TIT319_High"
   IOField "I/O field_115" at 1208,311 size 60x22; Authorization "Parameter Change"; FormatPattern s999.9
      ProcessValue <- "84_Setpoints_TIT319_HighHigh"
   IOField "I/O field_119" at 1140,351 size 60x22; Authorization "Parameter Change"; FormatPattern s999.9
      ProcessValue <- "84_Setpoints_TIT360_High"
   IOField "I/O field_120" at 1208,351 size 60x22; Authorization "Parameter Change"; FormatPattern s999.9
      ProcessValue <- "84_Setpoints_TIT360_HighHigh"
   IOField "I/O field_124" at 1140,391 size 60x22; Authorization "Parameter Change"; FormatPattern 99.9
      ProcessValue <- "84_Setpoints_PIT359_High"
   IOField "I/O field_125" at 1208,391 size 60x22; Authorization "Parameter Change"; FormatPattern 99.9
      ProcessValue <- "84_Setpoints_PIT359_HighHigh"
   IOField "I/O field_84" at 1139,431 size 60x22; Authorization "Parameter Change"; FormatPattern 99.9
      ProcessValue <- "84_Setpoints_PIT316_High"
   IOField "I/O field_85" at 1207,431 size 60x22; Authorization "Parameter Change"; FormatPattern 99.9
      ProcessValue <- "84_Setpoints_PIT316_HighHigh"
   IOField "I/O field_122" at 1004,391 size 60x22; Authorization "Parameter Change"; FormatPattern 99.9
      ProcessValue <- "84_Setpoints_PIT359_LowLow"
   IOField "I/O field_123" at 1072,391 size 60x22; Authorization "Parameter Change"; FormatPattern 99.9
      ProcessValue <- "84_Setpoints_PIT359_Low"
   IOField "I/O field_82" at 1003,431 size 60x22; Authorization "Parameter Change"; FormatPattern 99.9
      ProcessValue <- "84_Setpoints_PIT316_LowLow"
   IOField "I/O field_83" at 1071,431 size 60x22; Authorization "Parameter Change"; FormatPattern 99.9
      ProcessValue <- "84_Setpoints_PIT316_Low"
   TextField "Text field_52" at 17,91 size 340x26; Text 'BWT Control System PLC (Rack 3)'
   TextField "Text field_54" at 649,719 size 228x62; Text 'Note: CSW = Cooling Sea Water'
   Button "Button_1" at 1160,732 size 100x35; TextOn 'BWTS Digital Inputs.'; TextOff 'Next'
      on Click: ActivateScreen("BC Analogue Inputs", 0)
   TextField "Text field_25" at 60,231 size 220x22; Text 'PIT-102 - CA Pressure (Post-Ignition)'
   IOField "I/O field_52" at 361,231 size 60x22; Authorization "Parameter Change"; FormatPattern 9999
      ProcessValue <- "84_Setpoints_PIT102_Post_LowLow"
   IOField "I/O field_53" at 429,231 size 60x22; Authorization "Parameter Change"; FormatPattern 9999
      ProcessValue <- "84_Setpoints_PIT102_Post_Low"
   IOField "I/O field_54" at 497,231 size 60x22; Authorization "Parameter Change"; FormatPattern 9999
      ProcessValue <- "84_Setpoints_PIT102_Post_High"
   IOField "I/O field_55" at 565,231 size 60x22; Authorization "Parameter Change"; FormatPattern 9999
      ProcessValue <- "84_Setpoints_PIT102_Post_HighHigh"
   TextField "Text field_32" at 7,231 size 53x22; Text 'IW112'
   TextField "Text field_33" at 60,391 size 220x22; Text 'PIT-402 - IG Outlet Pres. (Post-Ignitn)'
   IOField "I/O field_57" at 361,391 size 60x22; Authorization "Parameter Change"; FormatPattern 9999
      ProcessValue <- "84_Setpoints_PIT402_Post_LowLow"
   IOField "I/O field_58" at 429,391 size 60x22; Authorization "Parameter Change"; FormatPattern 9999
      ProcessValue <- "84_Setpoints_PIT402_Post_Low"
   IOField "I/O field_59" at 497,391 size 60x22; Authorization "Parameter Change"; FormatPattern 9999
      ProcessValue <- "84_Setpoints_PIT402_Post_High"
   IOField "I/O field_60" at 565,391 size 60x22; Authorization "Parameter Change"; FormatPattern 9999
      ProcessValue <- "84_Setpoints_PIT402_Post_HighHigh"
   TextField "Text field_34" at 7,391 size 53x22; Text 'IW116'
   IOField "I/O field_47" at 1004,191 size 60x22; Authorization "Commissioning"; FormatPattern 99.9
      ProcessValue <- "84_Setpoints_AT_O2_2_LowLow"
   IOField "I/O field_48" at 1072,191 size 60x22; Authorization "Commissioning"; FormatPattern 99.9
      ProcessValue <- "84_Setpoints_AT_O2_2_Low"
   TextField "Text field_35" at 61,191 size 220x22; Text 'PIT-102 - CA Pressure (Main)'
   IOField "I/O field_50" at 362,191 size 60x22; Authorization "Parameter Change"; FormatPattern 9999
      ProcessValue <- "84_Setpoints_PIT102_Main_LowLow"
   IOField "I/O field_63" at 430,191 size 60x22; Authorization "Parameter Change"; FormatPattern 9999
      ProcessValue <- "84_Setpoints_PIT102_Main_Low"
   IOField "I/O field_64" at 498,191 size 60x22; Authorization "Parameter Change"; FormatPattern 9999
      ProcessValue <- "84_Setpoints_PIT102_Main_High"
   IOField "I/O field_65" at 566,191 size 60x22; Authorization "Parameter Change"; FormatPattern 9999
      ProcessValue <- "84_Setpoints_PIT102_Main_HighHigh"
   TextField "Text field_36" at 8,191 size 53x22; Text 'IW112'
   IOField "I/O field_49" at 1004,231 size 60x22; FormatPattern 999
   IOField "I/O field_51" at 1072,231 size 60x22; FormatPattern 999
   IOField "I/O field_66" at 1140,231 size 60x22; FormatPattern 999
   IOField "I/O field_67" at 1208,231 size 60x22; FormatPattern 999
   TextField "Text field_37" at 61,349 size 220x22; Text 'PIT-402 - IG Outlet Pres. (Main)'
   IOField "I/O field_69" at 362,349 size 60x22; Authorization "Parameter Change"; FormatPattern 9999
      ProcessValue <- "84_Setpoints_PIT402_Main_LowLow"
   IOField "I/O field_70" at 430,349 size 60x22; Authorization "Parameter Change"; FormatPattern 9999
      ProcessValue <- "84_Setpoints_PIT402_Main_Low"
   IOField "I/O field_71" at 498,349 size 60x22; Authorization "Parameter Change"; FormatPattern 9999
      ProcessValue <- "84_Setpoints_PIT402_Main_High"